screen "BC Process Times" 1280x800, template "Template"
   on GenerateScreen: "TitleUpdater"()
   Button "HmiScreenItemData_1" at 1,1 size 150x43; TextOn 'Back'; TextOff 'Commissioning'
      on Release: ActivateScreen("Commissioning Main Page", 0)
   Button "Button_1" at 21,736 size 161x32; TextOff 'IGG Step Times'
      on Activate: ActivateScreen("IGG Max Step Times", 0)
   Button "Button_2" at 1091,736 size 161x32; TextOff 'BC Step Times'
      on Activate: ActivateScreen("BC Max Step Times", 0)
   AlarmView "Alarm view_1" at 0,777 size 1280x23
   TextField "Text field_2" at 262,326 size 271x22; Text 'CV114 Open Delay Time'
   TextField "Text field_3" at 551,161 size 65x20; Text 'Time (s)'
   TextField "Text field_4" at 262,354 size 273x22; Text 'CV206 Open Delay Time'
   IOField "I/O field_1" at 546,354 size 60x22; Authorization "Parameter Change"; FormatPattern 999
      ProcessValue <- "86_Times_CV206_OPEN_TIME"
   TextField "Text field_5" at 262,411 size 270x22; Text 'CV215 Open Delay Time'
   TextField "Text field_6" at 262,186 size 272x22; Text 'CV127 Open #1 Delay Time'
   TextField "Text field_7" at 262,214 size 272x22; Text 'CV127 Closed Delay Time'
   TextField "Text field_8" at 262,242 size 271x22; Text 'CV127 Open #2 Delay Time'
   TextField "Text field_9" at 262,270 size 270x22; Text 'CV124 Open Delay Time'
   TextField "Text field_10" at 262,298 size 270x22; Text 'CV124 Close Delay Purge Time'
   TextField "Text field_11" at 262,161 size 89x20; Text 'Description'
   IOField "I/O field_3" at 546,186 size 60x22; Authorization "Parameter Change"; FormatPattern 999
      ProcessValue <- "86_Times_CV127_OPEN_TIME_#1"
   IOField "I/O field_4" at 546,214 size 60x22; Authorization "Parameter Change"; FormatPattern 999
      ProcessValue <- "86_Times_CV127_CLOSED_TIME"
   IOField "I/O field_6" at 546,242 size 60x22; Authorization "Parameter Change"; FormatPattern 999
      ProcessValue <- "86_Times_CV127_OPEN_TIME_#2"
   IOField "I/O field_8" at 546,298 size 60x22; Authorization "Parameter Change"; FormatPattern 999
      ProcessValue <- "86_Times_CV124_CLOSE_TIME_PRG"
   IOField "I/O field_9" at 546,410 size 60x22; Authorization "Parameter Change"; FormatPattern 999
      ProcessValue <- "86_Times_CV215_OPEN_TIME"
   TextField "Text field_12" at 261,135 size 178x26; Text 'BC Process Times'
   IOField "I/O field_10" at 546,270 size 60x22; Authorization "Parameter Change"; FormatPattern 999
      ProcessValue <- "86_Times_CV124_OPEN_TIME"
   TextField "Text field_13" at 262,383 size 270x22; Text 'CV207 Open Delay Time'
   IOField "I/O field_11" at 546,382 size 60x22; Authorization "Parameter Change"; FormatPattern 999
      ProcessValue <- "86_Times_CV207_OPEN_TIME"
   TextField "Text field_17" at 262,439 size 270x22; Text 'CV215 Close Delay Purge Time'
   IOField "I/O field_16" at 546,438 size 60x22; Authorization "Parameter Change"; FormatPattern 999
      ProcessValue <- "86_Times_CV215_CLOSE_TIME_PRG"
   TextField "Text field_18" at 262,467 size 270x22; Text 'CV216 Open Delay Time'
   IOField "I/O field_17" at 546,466 size 60x22; Authorization "Parameter Change"; FormatPattern 999
      ProcessValue <- "86_Times_CV216_OPEN_TIME"
   TextField "Text field_19" at 262,495 size 269x22; Text 'CV216 Close Delay Purge Time'
   IOField "I/O field_18" at 546,494 size 60x22; Authorization "Parameter Change"; FormatPattern 999
      ProcessValue <- "86_Times_CV216_CLOSE_TIME_PRG"
   TextField "Text field_20" at 262,523 size 269x22; Text 'CV216 Open Delay Purge Time'
   IOField "I/O field_19" at 546,522 size 60x22; Authorization "Parameter Change"; FormatPattern 999
      ProcessValue <- "86_Times_CV216_OPEN_TIME_PRG"
   TextField "Text field_21" at 262,552 size 269x22; Text 'CV206 Close Delay Time'
   IOField "I/O field_20" at 546,551 size 60x22; Authorization "Parameter Change"; FormatPattern 999
      ProcessValue <- "86_Times_CV206_CLOSE_TIME"
   TextField "Text field_22" at 636,186 size 269x22; Text 'CV207 Close Delay Time'
   IOField "I/O field_21" at 916,186 size 60x22; Authorization "Parameter Change"; FormatPattern 999
      ProcessValue <- "86_Times_CV207_CLOSE_TIME"
   TextField "Text field_23" at 636,160 size 89x20; Text 'Description'
   TextField "Text field_24" at 923,161 size 65x20; Text 'Time (s)'
   TextField "Text field_26" at 636,214 size 269x22; Text 'CV114 Close Delay Time'
   IOField "I/O field_22" at 916,214 size 60x22; Authorization "Parameter Change"; FormatPattern 999
      ProcessValue <- "86_Times_CV114_CLOSE_TIME"
   TextField "Text field_27" at 636,242 size 269x22; Text 'CV215 Close Delay Time'
   IOField "I/O field_23" at 916,242 size 60x22; Authorization "Parameter Change"; FormatPattern 999
      ProcessValue <- "86_Times_CV215_CLOSE_TIME"
   TextField "Text field_28" at 636,270 size 269x22; Text 'CV216 Close Delay Time'
   IOField "I/O field_24" at 916,270 size 60x22; Authorization "Parameter Change"; FormatPattern 999
      ProcessValue <- "86_Times_CV216_CLOSE_TIME"
   TextField "Text field_30" at 636,298 size 269x22; Text 'CV124 Close Delay Time'
   IOField "I/O field_25" at 916,298 size 60x22; Authorization "Parameter Change"; FormatPattern 999
      ProcessValue <- "86_Times_CV124_CLOSE_TIME"
   TextField "Text field_31" at 636,326 size 269x22; Text 'X001 Maximum Run Time'
   IOField "I/O field_26" at 916,326 size 60x22; Authorization "Parameter Change"; FormatPattern 999
      ProcessValue <- "86_Times_X001_MAX_RUN_TIME"
   TextField "Text field_32" at 636,354 size 269x22; Text 'X001 Run Confirmation Time'
   IOField "I/O field_27" at 916,354 size 60x22; Authorization "Parameter Change"; FormatPattern 999
      ProcessValue <- "86_Times_X001_RUN_CNF_TIME"
   TextField "Text field_34" at 636,383 size 269x22; Text 'Flame Detection Delay'
   IOField "I/O field_28" at 916,382 size 60x22; Authorization "Parameter Change"; FormatPattern 999
      ProcessValue <- "86_Times_FD_DET_DELAY"
   TextField "Text field_36" at 636,411 size 269x22; Text 'Flame Verification Time'
   IOField "I/O field_29" at 916,410 size 60x22; Authorization "Parameter Change"; FormatPattern 999
      ProcessValue <- "86_Times_FD_VRFCTN_TIME"
   TextField "Text field_37" at 636,439 size 269x22; Text 'Flame Detection Time'
   IOField "I/O field_30" at 916,438 size 60x22; Authorization "Parameter Change"; FormatPattern 999
      ProcessValue <- "86_Times_FDU_DET_TIME"
   TextField "Text field_38" at 636,467 size 269x22; Text 'Max Ignition Sequence Run Time'
   IOField "I/O field_31" at 916,466 size 60x22; Authorization "Parameter Change"; FormatPattern 999
      ProcessValue <- "86_Times_MAX_IGNTN_SEQ_TIME"
   TextField "Text field_39" at 636,495 size 269x22; Text 'Max Main Burner Sequence Run Time'
      Visibility <- "AlwaysTRUE"
   IOField "I/O field_32" at 916,494 size 60x22; Authorization "Parameter Change"; FormatPattern 999; Unit h
      Visibility <- "AlwaysTRUE"
      ProcessValue <- "86_Times_MAX_MAIN_BURN_SEQ_TIME"
   TextField "Text field_40" at 636,523 size 269x22; Text 'Max Pilot Burner Purge Sequence Run Time'
   IOField "I/O field_33" at 916,522 size 60x22; Authorization "Parameter Change"; FormatPattern 999
      ProcessValue <- "86_Times_MAX_PILOT_PURGE_SEQ_TIME"
   TextField "Text field_41" at 636,552 size 269x22; Text 'O2 Check Delay Time'
   IOField "I/O field_34" at 916,551 size 60x22; Authorization "Parameter Change"; FormatPattern 999
      ProcessValue <- "86_Times_O2_CHECK_TIME"
   IOField "I/O field_7" at 546,326 size 60x22; Authorization "Parameter Change"; FormatPattern 999
      ProcessValue <- "86_Times_CV114_OPEN_TIME"
   TextField "Text field_43" at 636,582 size 269x22; Text 'Flame Fail Delay'
   IOField "I/O field_35" at 916,581 size 60x22; Authorization "Parameter Change"; FormatPattern 999
      ProcessValue <- "80_From_HMI_FLM_FAIL_DLY"
   Switch "Switch_1" at 987,492 size 32x29; CaptionText 'Switch'; TextOn 'ON'; TextOff 'OFF'; Authorization "User administration"; PictureOff "Design_5_PilotLight_Green_Off"; PictureOn "Design_5_PilotLight_Green_On"
      on Activate: SetBit("80_From_HMI_BurnerProgramedStop")
      Visibility <- "AlwaysTRUE"
      ProcessValue <- "80_From_HMI_BurnerProgramedStop"
   TextField "Text field_44" at 636,613 size 269x22; Text 'FS317 Delayed Fault'
   IOField "I/O field_36" at 916,613 size 60x22; Authorization "Parameter Change"; FormatPattern 999
      ProcessValue <- "86_Times_FS317 delay"
   TextField "Text field_45" at 636,644 size 269x22; Text 'FS320 Delayed Fault'
   IOField "I/O field_37" at 916,644 size 60x22; Authorization "Parameter Change"; FormatPattern 999
      ProcessValue <- "86_Times_FS320 delay"
   TextField "Text field_46" at 262,581 size 269x22; Text 'FS359 Delayed Fault'
   IOField "I/O field_38" at 546,581 size 60x22; Authorization "Parameter Change"; FormatPattern 999
      ProcessValue <- "80_From_HMI_PIT 359 delay"
   TextField "Text field_47" at 262,612 size 269x22; Text 'FS316 Delayed Fault'
   IOField "I/O field_39" at 546,612 size 60x22; Authorization "Parameter Change"; FormatPattern 999
      ProcessValue <- "80_From_HMI_PIT 316 delay"
   Group "Group" at 455,41 size 373x50
   TextField "Text field_1" at 262,643 size 269x22; Text 'PS101 Delayed Fault'
   IOField "I/O field_2" at 546,643 size 60x22; Authorization "Parameter Change"; FormatPattern 999
      ProcessValue <- "86_Times_PS101 Alarm Delay"
   Button "HmiScreenItemData_8" at 469,45 size 355x40; TextOn 'Back'; TextOff 'Text'
   TextField "Screen title" at 455,41 size 373x50; Text 'Screen title'

screen "GCU Process Times" 1280x800, template "Template"
   on GenerateScreen: "TitleUpdater"()
   Button "HmiScreenItemData_1" at 1,1 size 150x43; TextOn 'Back'; TextOff 'Commissioning'
      on Release: ActivateScreen("Commissioning Main Page", 0)
   AlarmView "Alarm view_1" at 0,777 size 1280x23
   TextField "Text field_29" at 545,103 size 65x20; Text 'Time (s)'
   TextField "Text field_65" at 240,128 size 300x25; Text 'P303 Started Delay'
   TextField "Text field_42" at 240,103 size 89x20; Text 'Description'
   IOField "I/O field_128" at 545,128 size 65x25; Authorization "Parameter Change"; FormatPattern 999
      ProcessValue <- "86_Times_P303_STRTD_DLY"
   TextField "Text field_53" at 240,74 size 193x26; Text 'GCU Process Times'
   TextField "Text field_1" at 240,158 size 300x25; Text 'P303 Stopped Delay'
   IOField "I/O field_1" at 545,158 size 65x25; Authorization "Parameter Change"; FormatPattern 999
      ProcessValue <- "86_Times_P303_STPD_DLY"
   TextField "Text field_2" at 240,188 size 300x25; Text 'P304 Started Delay'
   IOField "I/O field_2" at 545,188 size 65x25; Authorization "Parameter Change"; FormatPattern 999
      ProcessValue <- "86_Times_P304_STRTD_DLY"
   TextField "Text field_3" at 240,218 size 300x25; Text 'P304 Stopped Delay'
   IOField "I/O field_3" at 545,218 size 65x25; Authorization "Parameter Change"; FormatPattern 999
      ProcessValue <- "86_Times_P304_STPD_DLY"
   TextField "Text field_4" at 240,248 size 300x25; Text 'P305 Started Delay'
   IOField "I/O field_4" at 545,248 size 65x25; Authorization "Parameter Change"; FormatPattern 999
      ProcessValue <- "86_Times_P305_STRTD_DLY"
   TextField "Text field_5" at 240,278 size 300x25; Text 'P305 Stopped Delay'
   IOField "I/O field_5" at 545,278 size 65x25; Authorization "Parameter Change"; FormatPattern 999
      ProcessValue <- "86_Times_P305_STPD_DLY"
   TextField "Text field_6" at 240,308 size 300x25; Text 'CV341 Closed Delay'
   IOField "I/O field_6" at 545,308 size 65x25; Authorization "Parameter Change"; FormatPattern 999
      ProcessValue <- "86_Times_CV341_CLSD_DLY"
   TextField "Text field_7" at 240,338 size 300x25; Text 'CV358 Closed Delay'
   IOField "I/O field_7" at 545,338 size 65x25; Authorization "Parameter Change"; FormatPattern 999
      ProcessValue <- "86_Times_CV358_CLSD_DLY"
   TextField "Text field_8" at 975,103 size 65x20; Text 'Time (s)'
   TextField "Text field_9" at 670,128 size 300x25; Text 'CV405 Opened Delay'
   TextField "Text field_10" at 670,103 size 89x20; Text 'Description'
   IOField "I/O field_8" at 975,128 size 65x25; Authorization "Parameter Change"; FormatPattern 999
      ProcessValue <- "86_Times_CV405_OPND_DLY"
   TextField "Text field_11" at 670,158 size 300x25; Text 'CV406 Closed Delay'
   IOField "I/O field_9" at 975,158 size 65x25; Authorization "Parameter Change"; FormatPattern 999
      ProcessValue <- "86_Times_CV406_CLSD_DLY"
   TextField "Text field_12" at 670,188 size 300x25; Text 'E400 Stop Time'
   IOField "I/O field_10" at 975,188 size 65x25; Authorization "Parameter Change"; FormatPattern 999
      ProcessValue <- "86_Times_E400_STOP_TIME"
   TextField "Text field_13" at 670,218 size 300x25; Text 'P303 Stop Time'
   IOField "I/O field_11" at 975,218 size 65x25; Authorization "Parameter Change"; FormatPattern 999
      ProcessValue <- "86_Times_P303_STOP_TIME"
   TextField "Text field_14" at 670,248 size 300x25; Text 'CV341 Opened Delay'
   IOField "I/O field_12" at 975,248 size 65x25; Authorization "Parameter Change"; FormatPattern 999
      ProcessValue <- "86_Times_CV341_OPND_DLY"
   TextField "Text field_15" at 670,278 size 300x25; Text 'GCU Tank Maximum Drain Time'
   IOField "I/O field_13" at 975,278 size 65x25; Authorization "Parameter Change"; FormatPattern 999
      ProcessValue <- "86_Times_GCU_TNK_DRN_MAX_TIME"
   TextField "Text field_16" at 670,308 size 300x25; Text 'GCU Flush Time'
   IOField "I/O field_14" at 975,308 size 65x25; Authorization "Parameter Change"; FormatPattern 999
      ProcessValue <- "86_Times_GCU_FLUSH_TIME"
   TextField "Text field_17" at 670,338 size 300x25; Text 'Post Flush Delay'
   IOField "I/O field_15" at 975,338 size 65x25; Authorization "Parameter Change"; FormatPattern 999
      ProcessValue <- "86_Times_POST_FLUSH_DLY"
   TextField "Text field_18" at 240,368 size 300x25; Text 'CV401 Opened Delay'
   IOField "I/O field_16" at 545,368 size 65x25; Authorization "Parameter Change"; FormatPattern 999
      ProcessValue <- "86_Times_CV401_OPND_DLY"
   TextField "Text field_19" at 240,398 size 300x25; Text 'CV401 Closed Delay'
   IOField "I/O field_17" at 545,398 size 65x25; Authorization "Parameter Change"; FormatPattern 999
      ProcessValue <- "86_Times_CV401_CLSD_DLY"
   TextField "Text field_20" at 240,428 size 300x25; Text 'CV441 Opened Delay'
   IOField "I/O field_18" at 545,428 size 65x25; Authorization "Parameter Change"; FormatPattern 999
      ProcessValue <- "86_Times_CV441_OPND_DLY"
   TextField "Text field_21" at 240,458 size 300x25; Text 'CV441 Closed Delay'
   IOField "I/O field_19" at 545,458 size 65x25; Authorization "Parameter Change"; FormatPattern 999
      ProcessValue <- "86_Times_CV441_CLSD_DLY"
   TextField "Text field_22" at 240,488 size 300x25; Text 'Pre CV441 Open Delay'
   IOField "I/O field_20" at 545,488 size 65x25; Authorization "Parameter Change"; FormatPattern 999
      ProcessValue <- "86_Times_PRE_CV441_OPN_DLY"
   TextField "Text field_23" at 240,518 size 300x25; Text 'Valve Configuration Done Delay'
   IOField "I/O field_21" at 545,518 size 65x25; Authorization "Parameter Change"; FormatPattern 999
      ProcessValue <- "86_Times_VLV_CNFG_DN_DLY"
   TextField "Text field_24" at 240,548 size 300x25; Text 'Pre GCU Tank Fill Delay'
   IOField "I/O field_22" at 545,548 size 65x25; Authorization "Parameter Change"; FormatPattern 999
      ProcessValue <- "86_Times_PRE_GCU_TNK_FILL_DLY"
   TextField "Text field_25" at 240,578 size 300x25; Text 'GCU Tank Fill Maximum Time'
   IOField "I/O field_23" at 545,578 size 65x25; Authorization "Parameter Change"; FormatPattern 999
      ProcessValue <- "86_Times_GCU_TNK_FILL_MAX_TIME"
   TextField "Text field_26" at 670,368 size 300x25; Text 'CV341 Maximum Travel Time'
   IOField "I/O field_24" at 975,368 size 65x25; Authorization "Parameter Change"; FormatPattern 999
      ProcessValue <- "86_Times_CV341_MAX_TRVL_TIME"
   TextField "Text field_27" at 670,398 size 300x25; Text 'CV358 Maximum Travel Time'
   IOField "I/O field_25" at 975,398 size 65x25; Authorization "Parameter Change"; FormatPattern 999
      ProcessValue <- "86_Times_CV358_MAX_TRVL_TIME"
   TextField "Text field_28" at 670,428 size 300x25; Text 'CV406 Maximum Travel Time'
   IOField "I/O field_26" at 975,428 size 65x25; Authorization "Parameter Change"; FormatPattern 999
      ProcessValue <- "86_Times_CV406_MAX_TRVL_TIME"
   TextField "Text field_30" at 670,458 size 300x25; Text 'CV407 Maximum Travel Time'
   IOField "I/O field_27" at 975,458 size 65x25; Authorization "Parameter Change"; FormatPattern 999
      ProcessValue <- "86_Times_CV407_MAX_TRVL_TIME"
   TextField "Text field_31" at 670,488 size 300x25; Text 'CV409 Maximum Travel Time'
   IOField "I/O field_28" at 975,488 size 65x25; Authorization "Parameter Change"; FormatPattern 999
      ProcessValue <- "86_Times_CV409_MAX_TRVL_TIME"
   TextField "Text field_32" at 670,518 size 300x25; Text 'CV411 Maximum Travel Time'
   IOField "I/O field_29" at 975,518 size 65x25; Authorization "Parameter Change"; FormatPattern 999
      ProcessValue <- "86_Times_CV411_MAX_TRVL_TIME"
   TextField "Text field_33" at 670,548 size 300x25; Text 'CV441 Maximum Travel Time'
   IOField "I/O field_30" at 975,548 size 65x25; Authorization "Parameter Change"; FormatPattern 999
      ProcessValue <- "86_Times_CV441_MAX_TRVL_TIME"
   TextField "Text field_34" at 670,638 size 300x25; Text 'PIT416 Target Ramp Time'
   IOField "I/O field_31" at 975,638 size 65x25; Authorization "Parameter Change"; FormatPattern 999
      ProcessValue <- "86_Times_PIT416_TRGT_RMP_TIME"
   TextField "Text field_35" at 240,608 size 300x25; Text 'E400 Started Delay'
   IOField "I/O field_32" at 545,608 size 65x25; Authorization "Parameter Change"; FormatPattern 999
      ProcessValue <- "86_Times_E400_STRTD_DLY"
   TextField "Text field_36" at 240,638 size 300x25; Text 'E400 Running Delay'
   IOField "I/O field_33" at 545,638 size 65x25; Authorization "Parameter Change"; FormatPattern 999
      ProcessValue <- "86_Times_E400_RNG_DLY"
   TextField "Text field_37" at 670,578 size 300x25; Text 'PIT353 Alarm Delay Time'
   IOField "I/O field_34" at 975,578 size 65x25; Authorization "Parameter Change"; FormatPattern 999
      ProcessValue <- "86_Times_PIT353 Delay"
   TextField "Text field_38" at 670,608 size 300x25; Text 'PIT416 Alarm Delay Time'
   IOField "I/O field_35" at 975,608 size 65x25; Authorization "Parameter Change"; FormatPattern 999
      ProcessValue <- "86_Times_PIT416 Delay"
   TextField "Text field_39" at 240,669 size 300x25; Text 'P301 Started Delay'
   IOField "I/O field_36" at 545,669 size 65x25; Authorization "Parameter Change"; FormatPattern 999
      ProcessValue <- "86_Times_P301_START_DLY"
   TextField "Text field_40" at 670,669 size 300x25; Text 'FS332 Alarm Delay'
   IOField "I/O field_37" at 975,669 size 65x25; Authorization "Parameter Change"; FormatPattern 999
      ProcessValue <- "86_Times_FS332 Delay"
   TextField "Text field_41" at 670,701 size 300x25; Text 'LIT304 Alarm Delay'
   IOField "I/O field_38" at 975,701 size 65x25; Authorization "Parameter Change"; FormatPattern 999
      ProcessValue <- "86_Times_LIT304 Delay"
   Group "Group" at 455,41 size 373x50
   TextField "Text field_43" at 240,701 size 300x25; Text 'PIT358 Alarm Delay Time'
   IOField "I/O field_39" at 545,701 size 65x25; Authorization "Parameter Change"; FormatPattern 999
      ProcessValue <- "86_Times_PIT358 Delay"
   TextField "Text field_44" at 240,732 size 300x25; Text 'PIT348 Alarm Delay Time'
   IOField "I/O field_40" at 545,732 size 65x25; Authorization "Parameter Change"; FormatPattern 999
      ProcessValue <- "86_Times_PIT348 Delay"
   Button "HmiScreenItemData_8" at 469,45 size 355x40; TextOn 'Back'; TextOff 'Text'
   TextField "Screen title" at 455,41 size 373x50; Text 'Screen title'

screen "GCU Max Step Times" 1280x800, template "Template"
   on GenerateScreen: "TitleUpdater"()
   Button "HmiScreenItemData_1" at 1,1 size 150x43; TextOn 'Back'; TextOff 'Commissioning'
      on Release: ActivateScreen("Commissioning Main Page", 0)
   TextField "Text field_29" at 130,95 size 75x25; Text 'Time (ms)'
   TextField "Text field_65" at 40,130 size 75x25; Text 'Step 001'
   TextField "Text field_42" at 40,95 size 75x25; Text 'STEP'
   IOField "I/O field_128" at 130,130 size 75x25; Authorization "Parameter Change"; FormatPattern 999999
      ProcessValue <- "86_Times_STEP_MAX_TIME_STP_001"
   TextField "Text field_53" at 40,66 size 262x26; Text 'GCU Maximum Step Times'
   TextField "Text field_1" at 385,95 size 75x25; Text 'Time (ms)'
   TextField "Text field_2" at 295,130 size 75x25; Text 'Step 170'
   TextField "Text field_3" at 295,95 size 75x25; Text 'STEP'
   IOField "I/O field_1" at 385,130 size 75x25; Authorization "Parameter Change"; FormatPattern 999999
      ProcessValue <- "86_Times_STEP_MAX_TIME_STP_170"
   TextField "Text field_4" at 640,95 size 75x25; Text 'Time (ms)'
   TextField "Text field_5" at 550,130 size 75x25; Text 'Step 350'
   TextField "Text field_6" at 550,95 size 75x25; Text 'STEP'
   IOField "I/O field_2" at 640,130 size 75x25; Authorization "Parameter Change"; FormatPattern 999999
      ProcessValue <- "86_Times_STEP_MAX_TIME_STP_350"
   TextField "Text field_7" at 895,95 size 75x25; Text 'Time (ms)'
   TextField "Text field_8" at 805,130 size 75x25; Text 'Step 530'
   TextField "Text field_9" at 805,95 size 75x25; Text 'STEP'
   IOField "I/O field_3" at 895,130 size 75x25; Authorization "Parameter Change"; FormatPattern 999999
      ProcessValue <- "86_Times_STEP_MAX_TIME_STP_530"
   TextField "Text field_10" at 1150,95 size 75x25; Text 'Time (ms)'
   TextField "Text field_12" at 1060,95 size 75x25; Text 'STEP'
   TextField "Text field_13" at 40,165 size 75x25; Text 'Step 005'
   IOField "I/O field_5" at 130,165 size 75x25; Authorization "Parameter Change"; FormatPattern 999999
      ProcessValue <- "86_Times_STEP_MAX_TIME_STP_005"
   TextField "Text field_14" at 295,165 size 75x25; Text 'Step 180'
   IOField "I/O field_6" at 385,165 size 75x25; Authorization "Parameter Change"; FormatPattern 999999
      ProcessValue <- "86_Times_STEP_MAX_TIME_STP_180"
   TextField "Text field_15" at 550,165 size 75x25; Text 'Step 360'
   IOField "I/O field_7" at 640,165 size 75x25; Authorization "Parameter Change"; FormatPattern 999999
      ProcessValue <- "86_Times_STEP_MAX_TIME_STP_360"
   TextField "Text field_16" at 805,165 size 75x25; Text 'Step 540'
   IOField "I/O field_8" at 895,165 size 75x25; Authorization "Parameter Change"; FormatPattern 999999
      ProcessValue <- "86_Times_STEP_MAX_TIME_STP_540"
   TextField "Text field_18" at 40,200 size 75x25; Text 'Step 010'
   IOField "I/O field_10" at 130,200 size 75x25; Authorization "Parameter Change"; FormatPattern 999999
      ProcessValue <- "86_Times_STEP_MAX_TIME_STP_010"
   TextField "Text field_19" at 295,200 size 75x25; Text 'Step 190'
   IOField "I/O field_11" at 385,200 size 75x25; Authorization "Parameter Change"; FormatPattern 999999
      ProcessValue <- "86_Times_STEP_MAX_TIME_STP_190"
   TextField "Text field_20" at 550,200 size 75x25; Text 'Step 370'
   IOField "I/O field_12" at 640,200 size 75x25; Authorization "Parameter Change"; FormatPattern 999999
      ProcessValue <- "86_Times_STEP_MAX_TIME_STP_370"
   TextField "Text field_21" at 805,200 size 75x25; Text 'Step 550'
   IOField "I/O field_13" at 895,200 size 75x25; Authorization "Parameter Change"; FormatPattern 999999
      ProcessValue <- "86_Times_STEP_MAX_TIME_STP_550"
   TextField "Text field_23" at 40,235 size 75x25; Text 'Step 020'
   IOField "I/O field_15" at 130,235 size 75x25; Authorization "Parameter Change"; FormatPattern 999999
      ProcessValue <- "86_Times_STEP_MAX_TIME_STP_020"
   TextField "Text field_24" at 295,235 size 75x25; Text 'Step 200'
   IOField "I/O field_16" at 385,235 size 75x25; Authorization "Parameter Change"; FormatPattern 999999
      ProcessValue <- "86_Times_STEP_MAX_TIME_STP_200"
   TextField "Text field_25" at 550,235 size 75x25; Text 'Step 380'
   IOField "I/O field_17" at 640,235 size 75x25; Authorization "Parameter Change"; FormatPattern 999999
      ProcessValue <- "86_Times_STEP_MAX_TIME_STP_380"
   TextField "Text field_26" at 805,235 size 75x25; Text 'Step 560'
   IOField "I/O field_18" at 895,235 size 75x25; Authorization "Parameter Change"; FormatPattern 999999
      ProcessValue <- "86_Times_STEP_MAX_TIME_STP_560"
   TextField "Text field_28" at 40,270 size 75x25; Text 'Step 030'
   IOField "I/O field_20" at 130,270 size 75x25; Authorization "Parameter Change"; FormatPattern 999999
      ProcessValue <- "86_Times_STEP_MAX_TIME_STP_030"
   TextField "Text field_30" at 295,270 size 75x25; Text 'Step 210'
   IOField "I/O field_21" at 385,270 size 75x25; Authorization "Parameter Change"; FormatPattern 999999
      ProcessValue <- "86_Times_STEP_MAX_TIME_STP_210"
   TextField "Text field_31" at 550,270 size 75x25; Text 'Step 390'
   IOField "I/O field_22" at 640,270 size 75x25; Authorization "Parameter Change"; FormatPattern 999999
      ProcessValue <- "86_Times_STEP_MAX_TIME_STP_390"
   TextField "Text field_32" at 805,270 size 75x25; Text 'Step 570'
   IOField "I/O field_23" at 895,270 size 75x25; Authorization "Parameter Change"; FormatPattern 999999
      ProcessValue <- "86_Times_STEP_MAX_TIME_STP_570"
   TextField "Text field_34" at 40,305 size 75x25; Text 'Step 040'
   IOField "I/O field_25" at 130,305 size 75x25; Authorization "Parameter Change"; FormatPattern 999999
      ProcessValue <- "86_Times_STEP_MAX_TIME_STP_040"
   TextField "Text field_35" at 295,305 size 75x25; Text 'Step 220'
   IOField "I/O field_26" at 385,305 size 75x25; Authorization "Parameter Change"; FormatPattern 999999
      ProcessValue <- "86_Times_STEP_MAX_TIME_STP_220"
   TextField "Text field_36" at 550,305 size 75x25; Text 'Step 400'
   IOField "I/O field_27" at 640,305 size 75x25; Authorization "Parameter Change"; FormatPattern 999999
      ProcessValue <- "86_Times_STEP_MAX_TIME_STP_400"
   TextField "Text field_37" at 805,305 size 75x25; Text 'Step 580'
   IOField "I/O field_28" at 895,305 size 75x25; Authorization "Parameter Change"; FormatPattern 999999
      ProcessValue <- "86_Times_STEP_MAX_TIME_STP_580"
   TextField "Text field_39" at 40,340 size 75x25; Text 'Step 050'
   IOField "I/O field_30" at 130,340 size 75x25; Authorization "Parameter Change"; FormatPattern 999999
      ProcessValue <- "86_Times_STEP_MAX_TIME_STP_050"
   TextField "Text field_40" at 295,340 size 75x25; Text 'Step 230'
   IOField "I/O field_31" at 385,340 size 75x25; Authorization "Parameter Change"; FormatPattern 999999
      ProcessValue <- "86_Times_STEP_MAX_TIME_STP_230"
   TextField "Text field_41" at 550,340 size 75x25; Text 'Step 410'
   IOField "I/O field_32" at 640,340 size 75x25; Authorization "Parameter Change"; FormatPattern 999999
      ProcessValue <- "86_Times_STEP_MAX_TIME_STP_410"
   TextField "Text field_43" at 805,340 size 75x25; Text 'Step 590'
   IOField "I/O field_33" at 895,340 size 75x25; Authorization "Parameter Change"; FormatPattern 999999
      ProcessValue <- "86_Times_STEP_MAX_TIME_STP_590"
   TextField "Text field_45" at 40,375 size 75x25; Text 'Step 060'
   IOField "I/O field_35" at 130,375 size 75x25; Authorization "Parameter Change"; FormatPattern 999999
      ProcessValue <- "86_Times_STEP_MAX_TIME_STP_060"
   TextField "Text field_46" at 295,375 size 75x25; Text 'Step 240'
   IOField "I/O field_36" at 385,375 size 75x25; Authorization "Parameter Change"; FormatPattern 999999
      ProcessValue <- "86_Times_STEP_MAX_TIME_STP_240"
   TextField "Text field_47" at 550,375 size 75x25; Text 'Step 420'
   IOField "I/O field_37" at 640,375 size 75x25; Authorization "Parameter Change"; FormatPattern 999999
      ProcessValue <- "86_Times_STEP_MAX_TIME_STP_420"
   TextField "Text field_48" at 805,375 size 75x25; Text 'Step 600'
   IOField "I/O field_38" at 895,375 size 75x25; Authorization "Parameter Change"; FormatPattern 999999
      ProcessValue <- "86_Times_STEP_MAX_TIME_STP_600"
   TextField "Text field_50" at 40,410 size 75x25; Text 'Step 070'
   IOField "I/O field_40" at 130,410 size 75x25; Authorization "Parameter Change"; FormatPattern 999999
      ProcessValue <- "86_Times_STEP_MAX_TIME_STP_070"
   TextField "Text field_51" at 295,410 size 75x25; Text 'Step 250'
   IOField "I/O field_41" at 385,410 size 75x25; Authorization "Parameter Change"; FormatPattern 999999
      ProcessValue <- "86_Times_STEP_MAX_TIME_STP_250"
   TextField "Text field_52" at 550,410 size 75x25; Text 'Step 430'
   IOField "I/O field_42" at 640,410 size 75x25; Authorization "Parameter Change"; FormatPattern 999999
      ProcessValue <- "86_Times_STEP_MAX_TIME_STP_430"
   TextField "Text field_54" at 805,410 size 75x25; Text 'Step 610'
   IOField "I/O field_43" at 895,410 size 75x25; Authorization "Parameter Change"; FormatPattern 999999
      ProcessValue <- "86_Times_STEP_MAX_TIME_STP_610"
   TextField "Text field_56" at 40,445 size 75x25; Text 'Step 080'
   IOField "I/O field_45" at 130,445 size 75x25; Authorization "Parameter Change"; FormatPattern 999999
      ProcessValue <- "86_Times_STEP_MAX_TIME_STP_080"
   TextField "Text field_57" at 295,445 size 75x25; Text 'Step 260'
   IOField "I/O field_46" at 385,445 size 75x25; Authorization "Parameter Change"; FormatPattern 999999
      ProcessValue <- "86_Times_STEP_MAX_TIME_STP_260"
   TextField "Text field_58" at 550,445 size 75x25; Text 'Step 440'
   IOField "I/O field_47" at 640,445 size 75x25; Authorization "Parameter Change"; FormatPattern 999999
      ProcessValue <- "86_Times_STEP_MAX_TIME_STP_440"
   TextField "Text field_59" at 805,445 size 75x25; Text 'Step 620'
   IOField "I/O field_48" at 895,445 size 75x25; Authorization "Parameter Change"; FormatPattern 999999
      ProcessValue <- "86_Times_STEP_MAX_TIME_STP_620"
   TextField "Text field_61" at 40,480 size 75x25; Text 'Step 090'
   IOField "I/O field_50" at 130,480 size 75x25; Authorization "Parameter Change"; FormatPattern 999999
      ProcessValue <- "86_Times_STEP_MAX_TIME_STP_090"
   TextField "Text field_62" at 295,480 size 75x25; Text 'Step 270'
   IOField "I/O field_51" at 385,480 size 75x25; Authorization "Parameter Change"; FormatPattern 999999
      ProcessValue <- "86_Times_STEP_MAX_TIME_STP_270"
   TextField "Text field_63" at 550,480 size 75x25; Text 'Step 450'
   IOField "I/O field_52" at 640,480 size 75x25; Authorization "Parameter Change"; FormatPattern 999999
      ProcessValue <- "86_Times_STEP_MAX_TIME_STP_450"
   TextField "Text field_64" at 805,480 size 75x25; Text 'Step 630'
   IOField "I/O field_53" at 895,480 size 75x25; Authorization "Parameter Change"; FormatPattern 999999
      ProcessValue <- "86_Times_STEP_MAX_TIME_STP_630"
   TextField "Text field_67" at 40,515 size 75x25; Text 'Step 100'
   IOField "I/O field_55" at 130,515 size 75x25; Authorization "Parameter Change"; FormatPattern 999999
      ProcessValue <- "86_Times_STEP_MAX_TIME_STP_100"
   TextField "Text field_68" at 295,515 size 75x25; Text 'Step 280'
   IOField "I/O field_56" at 385,515 size 75x25; Authorization "Parameter Change"; FormatPattern 999999
      ProcessValue <- "86_Times_STEP_MAX_TIME_STP_280"
   TextField "Text field_69" at 550,515 size 75x25; Text 'Step 460'
   IOField "I/O field_57" at 640,515 size 75x25; Authorization "Parameter Change"; FormatPattern 999999
      ProcessValue <- "86_Times_STEP_MAX_TIME_STP_460"
   TextField "Text field_72" at 40,550 size 75x25; Text 'Step 110'
   IOField "I/O field_60" at 130,550 size 75x25; Authorization "Parameter Change"; FormatPattern 999999
      ProcessValue <- "86_Times_STEP_MAX_TIME_STP_110"
   TextField "Text field_73" at 295,550 size 75x25; Text 'Step 290'
   IOField "I/O field_61" at 385,550 size 75x25; Authorization "Parameter Change"; FormatPattern 999999
      ProcessValue <- "86_Times_STEP_MAX_TIME_STP_290"
   TextField "Text field_74" at 550,550 size 75x25; Text 'Step 470'
   IOField "I/O field_62" at 640,550 size 75x25; Authorization "Parameter Change"; FormatPattern 999999
      ProcessValue <- "86_Times_STEP_MAX_TIME_STP_470"
   TextField "Text field_77" at 40,585 size 75x25; Text 'Step 120'
   IOField "I/O field_65" at 130,585 size 75x25; Authorization "Parameter Change"; FormatPattern 999999
      ProcessValue <- "86_Times_STEP_MAX_TIME_STP_120"
   TextField "Text field_78" at 295,585 size 75x25; Text 'Step 300'
   IOField "I/O field_66" at 385,585 size 75x25; Authorization "Parameter Change"; FormatPattern 999999
      ProcessValue <- "86_Times_STEP_MAX_TIME_STP_300"
   TextField "Text field_79" at 550,585 size 75x25; Text 'Step 480'
   IOField "I/O field_67" at 640,585 size 75x25; Authorization "Parameter Change"; FormatPattern 999999
      ProcessValue <- "86_Times_STEP_MAX_TIME_STP_480"
   TextField "Text field_82" at 40,620 size 75x25; Text 'Step 130'
   IOField "I/O field_70" at 130,620 size 75x25; Authorization "Parameter Change"; FormatPattern 999999
      ProcessValue <- "86_Times_STEP_MAX_TIME_STP_130"
   TextField "Text field_83" at 295,620 size 75x25; Text 'Step 310'
   IOField "I/O field_71" at 385,620 size 75x25; Authorization "Parameter Change"; FormatPattern 999999
      ProcessValue <- "86_Times_STEP_MAX_TIME_STP_310"
   TextField "Text field_84" at 550,620 size 75x25; Text 'Step 490'
   IOField "I/O field_72" at 640,620 size 75x25; Authorization "Parameter Change"; FormatPattern 999999
      ProcessValue <- "86_Times_STEP_MAX_TIME_STP_490"
   TextField "Text field_87" at 40,655 size 75x25; Text 'Step 140'
   IOField "I/O field_75" at 130,655 size 75x25; Authorization "Parameter Change"; FormatPattern 999999
      ProcessValue <- "86_Times_STEP_MAX_TIME_STP_140"
   TextField "Text field_88" at 295,655 size 75x25; Text 'Step 320'
   IOField "I/O field_76" at 385,655 size 75x25; Authorization "Parameter Change"; FormatPattern 999999
      ProcessValue <- "86_Times_STEP_MAX_TIME_STP_320"
   TextField "Text field_89" at 550,655 size 75x25; Text 'Step 500'
   IOField "I/O field_77" at 640,655 size 75x25; Authorization "Parameter Change"; FormatPattern 999999
      ProcessValue <- "86_Times_STEP_MAX_TIME_STP_500"
   TextField "Text field_92" at 40,690 size 75x25; Text 'Step 150'
   IOField "I/O field_80" at 130,690 size 75x25; Authorization "Parameter Change"; FormatPattern 999999
      ProcessValue <- "86_Times_STEP_MAX_TIME_STP_150"
   TextField "Text field_93" at 295,690 size 75x25; Text 'Step 330'
   IOField "I/O field_81" at 385,690 size 75x25; Authorization "Parameter Change"; FormatPattern 999999
      ProcessValue <- "86_Times_STEP_MAX_TIME_STP_330"
   TextField "Text field_94" at 550,690 size 75x25; Text 'Step 510'
   IOField "I/O field_82" at 640,690 size 75x25; Authorization "Parameter Change"; FormatPattern 999999
      ProcessValue <- "86_Times_STEP_MAX_TIME_STP_510"
   TextField "Text field_97" at 40,725 size 75x25; Text 'Step 160'
   IOField "I/O field_85" at 130,725 size 75x25; Authorization "Parameter Change"; FormatPattern 999999
      ProcessValue <- "86_Times_STEP_MAX_TIME_STP_160"
   TextField "Text field_98" at 295,725 size 75x25; Text 'Step 340'
   IOField "I/O field_86" at 385,725 size 75x25; Authorization "Parameter Change"; FormatPattern 999999
      ProcessValue <- "86_Times_STEP_MAX_TIME_STP_340"
   TextField "Text field_99" at 550,725 size 75x25; Text 'Step 520'
   IOField "I/O field_87" at 640,725 size 75x25; Authorization "Parameter Change"; FormatPattern 999999
      ProcessValue <- "86_Times_STEP_MAX_TIME_STP_520"
   Group "Group" at 455,41 size 373x50
   Button "HmiScreenItemData_8" at 469,45 size 355x40; TextOn 'Back'; TextOff 'Text'
   TextField "Screen title" at 455,41 size 373x50; Text 'Screen title'

screen "GCU Target Setpoints" 1280x800, template "Template"
   on GenerateScreen: "TitleUpdater"()
   Button "HmiScreenItemData_1" at 1,1 size 150x43; TextOn 'Back'; TextOff 'Commissioning'
      on Release: ActivateScreen("Commissioning Main Page", 0)
   AlarmView "Alarm view_1" at 0,777 size 1280x23
   TextField "Text field_37" at 20,239 size 300x30; Text 'GCU Control PLC (Rack 3)'
   TextField "Text field_1" at 810,239 size 450x30; Text 'PROCESS STEP RELATED SETPOINTS & TARGETS'
   TextField "Text field_82" at 100,299 size 220x22; Text 'LIT304 GCU LEVEL'
   IOField "I/O field_22" at 350,299 size 70x22; FormatPattern 999; Unit  %
      ProcessValue <- "12_AI_Data_LIT_304_SCALED"
   IOField "I/O field_23" at 450,299 size 75x22; Authorization "Parameter Change"; FormatPattern 999
      ProcessValue <- "84_Setpoints_LIT304_InitialFill_LowLow"
   IOField "I/O field_24" at 550,299 size 75x22; Authorization "Parameter Change"; FormatPattern 999
      ProcessValue <- "84_Setpoints_LIT304_InitialFill_Low"
   IOField "I/O field_25" at 952,299 size 75x22; Authorization "Parameter Change"; FormatPattern 999
      ProcessValue <- "84_Setpoints_LIT304_InitialFill_High"
   IOField "I/O field_26" at 1052,299 size 75x22; Authorization "Parameter Change"; FormatPattern 999
      ProcessValue <- "84_Setpoints_LIT304_InitialFill_HighHigh"
   TextField "Text field_22" at 20,299 size 53x22; Text 'IW800'
   TextField "Text field_90" at 350,272 size 70x22; Text 'Reading'
   TextField "Text field_23" at 450,272 size 75x22; Text 'Low Low'
   TextField "Text field_26" at 550,272 size 75x22; Text 'Low'
   TextField "Text field_27" at 952,272 size 75x22; Text 'High'
   TextField "Text field_28" at 1052,272 size 75x22; Text 'High High'
   TextField "Text field_41" at 100,272 size 220x22; Text 'Description'
   TextField "Text field_43" at 20,272 size 53x22; Text 'AI'
   IOField "I/O field_27" at 750,299 size 75x22; Authorization "Parameter Change"; FormatPattern 999
      ProcessValue <- "84_Setpoints_LIT304_InitialFill_Target"
   TextField "Text field_29" at 750,272 size 75x22; Text 'Target'
   TextField "Text field_30" at 1152,299 size 100x22; Text 'INITIAL FILL'
   IOField "I/O field_28" at 450,339 size 75x22; Authorization "Parameter Change"; FormatPattern 999
      ProcessValue <- "84_Setpoints_LIT304_Refill_LowLow"
   IOField "I/O field_29" at 550,339 size 75x22; Authorization "Parameter Change"; FormatPattern 999
      ProcessValue <- "84_Setpoints_LIT304_Refill_Low"
   IOField "I/O field_30" at 952,339 size 75x22; Authorization "Parameter Change"; FormatPattern 999
      ProcessValue <- "84_Setpoints_LIT304_Refill_High"
   IOField "I/O field_40" at 1052,339 size 75x22; Authorization "Parameter Change"; FormatPattern 999
      ProcessValue <- "84_Setpoints_LIT304_Refill_HighHigh"
   IOField "I/O field_43" at 650,339 size 75x22; Authorization "Parameter Change"; FormatPattern 999
      ProcessValue <- "84_Setpoints_LIT304_Refill_Target_Low"
   TextField "Text field_31" at 1152,339 size 100x22; Text 'RE-FILL'
   IOField "I/O field_44" at 650,299 size 75x22; Authorization "Parameter Change"; FormatPattern 999
      ProcessValue <- "84_Setpoints_LIT304_InitialFill_Target_Low"
   TextField "Text field_32" at 645,272 size 83x22; Text 'Target Low'
   IOField "I/O field_45" at 750,339 size 75x22; Authorization "Parameter Change"; FormatPattern 999
      ProcessValue <- "84_Setpoints_LIT304_Refill_Target"
   TextField "Text field_2" at 100,379 size 220x22; Text 'PIT416 GAS TO DECK PRESS'
   IOField "I/O field_1" at 350,379 size 70x22; FormatPattern 9.9; Unit  Barg
      ProcessValue <- "12_AI_Data_PIT_416_SCALED"
   TextField "Text field_6" at 20,379 size 53x22; Text 'IW810'
   IOField "I/O field_4" at 750,379 size 75x22; Authorization "Parameter Change"; FormatPattern 9.9; Unit  Barg
      ProcessValue <- "84_Setpoints_PIT416_Target"
   TextField "Text field_7" at 100,419 size 220x22; Text 'PIT358 FCW INLET PRESS'
   IOField "I/O field_2" at 350,419 size 70x22; FormatPattern 9.9; Unit  Barg
      ProcessValue <- "12_AI_Data_PIT_358_SCALED"
   IOField "I/O field_3" at 450,419 size 75x22; Authorization "Parameter Change"; FormatPattern 9.9; Unit  Barg
      ProcessValue <- "84_Setpoints_PIT358_InitialFill_LowLow"
   IOField "I/O field_5" at 550,419 size 75x22; Authorization "Parameter Change"; FormatPattern 9.9; Unit  Barg
      ProcessValue <- "84_Setpoints_PIT358_InitialFill_Low"
   IOField "I/O field_6" at 952,419 size 75x22; Authorization "Parameter Change"; FormatPattern 99.9; Unit  Barg
      ProcessValue <- "84_Setpoints_PIT358_InitialFill_High"
   IOField "I/O field_7" at 1052,419 size 75x22; Authorization "Parameter Change"; FormatPattern 99.9; Unit  Barg
      ProcessValue <- "84_Setpoints_PIT358_InitialFill_HighHigh"
   TextField "Text field_8" at 20,419 size 53x22; Text 'IW812'
   TextField "Text field_9" at 1152,419 size 100x22; Text 'INITIAL FILL'
   IOField "I/O field_8" at 450,459 size 75x22; Authorization "Parameter Change"; FormatPattern 9.9; Unit  Barg
      ProcessValue <- "84_Setpoints_PIT358_Refill_LowLow"
   IOField "I/O field_9" at 550,459 size 75x22; Authorization "Parameter Change"; FormatPattern 9.9; Unit  Barg
      ProcessValue <- "84_Setpoints_PIT358_Refill_Low"
   IOField "I/O field_10" at 952,459 size 75x22; Authorization "Parameter Change"; FormatPattern 99.9; Unit  Barg
      ProcessValue <- "84_Setpoints_PIT358_Refill_High"
   IOField "I/O field_11" at 1052,459 size 75x22; Authorization "Parameter Change"; FormatPattern 99.9; Unit  Barg
      ProcessValue <- "84_Setpoints_PIT358_Refill_HighHigh"
   TextField "Text field_10" at 1152,459 size 100x22; Text 'RE-FILL'
   TextField "Text field_3" at 100,499 size 220x22; Text 'PIT353 RECIRC FCW PRESS'
   IOField "I/O field_12" at 350,499 size 70x22; FormatPattern 9.9; Unit  Barg
      ProcessValue <- "12_AI_Data_PIT_353_SCALED"
   IOField "I/O field_13" at 450,499 size 75x22; Authorization "Parameter Change"; FormatPattern 9.9; Unit  Barg
      ProcessValue <- "84_Setpoints_PIT353_InitialFill_LowLow"
   IOField "I/O field_14" at 550,499 size 75x22; Authorization "Parameter Change"; FormatPattern 9.9; Unit  Barg
      ProcessValue <- "84_Setpoints_PIT353_InitialFill_Low"
   IOField "I/O field_15" at 952,499 size 75x22; Authorization "Parameter Change"; FormatPattern 9.9; Unit  Barg
      ProcessValue <- "84_Setpoints_PIT353_InitialFill_High"
   IOField "I/O field_20" at 1052,499 size 75x22; Authorization "Parameter Change"; FormatPattern 9.9; Unit  Barg
      ProcessValue <- "84_Setpoints_PIT353_InitialFill_HighHigh"
   TextField "Text field_4" at 20,499 size 53x22; Text 'IW816'
   TextField "Text field_11" at 1152,499 size 100x22; Text 'INITIAL FILL'
   IOField "I/O field_21" at 450,539 size 75x22; Authorization "Parameter Change"; FormatPattern 9.9; Unit  Barg
      ProcessValue <- "84_Setpoints_PIT353_Refill_LowLow"
   IOField "I/O field_31" at 550,539 size 75x22; Authorization "Parameter Change"; FormatPattern 9.9; Unit  Barg
      ProcessValue <- "84_Setpoints_PIT353_Refill_Low"
   IOField "I/O field_32" at 952,539 size 75x22; Authorization "Parameter Change"; FormatPattern 9.9; Unit  Barg
      ProcessValue <- "84_Setpoints_PIT353_Refill_High"
   IOField "I/O field_33" at 1052,539 size 75x22; Authorization "Parameter Change"; FormatPattern 9.9; Unit  Barg
      ProcessValue <- "84_Setpoints_PIT353_Refill_HighHigh"
   TextField "Text field_12" at 1152,539 size 100x22; Text 'RE-FILL'
   TextField "Text field_5" at 836,272 size 107x22; Text 'Safe Target'
   IOField "I/O field_16" at 854,379 size 75x22; Authorization "Parameter Change"; FormatPattern 9.99; Unit  Barg
      ProcessValue <- "84_Setpoints_PIT416_Target_Safe"
   Group "Group" at 455,41 size 373x50
   Button "HmiScreenItemData_8" at 469,45 size 355x40; TextOn 'Back'; TextOff 'Text'
   TextField "Screen title" at 455,41 size 373x50; Text 'Screen title'

screen "Commissioning Main Page" 1280x800, template "Template"
   on GenerateScreen: "TitleUpdater"()
   Button "HmiScreenItemData_1" at 1,1 size 150x43; TextOn 'Back'; TextOff 'Main Index'
      on Release: ActivateScreen("02 Main Index", 0)
   AlarmView "Alarm view_1" at 0,777 size 1280x23
   Button "HmiScreenItemData_4" at 790,100 size 200x35; TextOn 'Back'; TextOff 'BWT Settings'
   Button "Button_22" at 800,150 size 180x50; TextOff 'Target Setpoints'; Authorization "Commissioning"
      on Press: ActivateScreen("BWT Target Setpoints", 0)
   Button "Button_24" at 800,220 size 180x50; TextOff 'Process Times'; Authorization "Commissioning"
      on Press: ActivateScreen("BWT Process Times", 0)
   Button "HmiScreenItemData_3" at 540,100 size 200x35; TextOn 'Back'; TextOff 'GCU Settings'
   Button "Button_13" at 550,150 size 180x50; TextOff 'Digital Inputs'; Authorization "Commissioning"
      on Click: ActivateScreen("GCU Digital Inputs", 0)
   Button "Button_14" at 550,220 size 180x50; TextOff 'Digital Outputs'; Authorization "Operating Mode"
      on Click: ActivateScreen("GCU Digital Outputs", 0)
   Button "Button_15" at 550,290 size 180x50; TextOff 'Analogue Inputs'; Authorization "Commissioning"
      on Press: ActivateScreen("GCU Analogue Inputs", 0)
   Button "Button_16" at 550,430 size 180x50; TextOff 'Target Setpoints'; Authorization "Commissioning"
      on Press: ActivateScreen("GCU Target Setpoints", 0)
   Button "Button_17" at 550,360 size 180x50; TextOff 'Analogue Outputs'; Authorization "Commissioning"
      on Press: ActivateScreen("GCU Analogue Outputs", 0)
   Button "Button_18" at 550,500 size 180x50; TextOff 'Process Times'; Authorization "Commissioning"
      on Press: ActivateScreen("GCU Process Times", 0)
   Button "HmiScreenItemData_2" at 290,100 size 200x35; TextOn 'Back'; TextOff 'IGG Settings'
   Button "Button_7" at 300,150 size 180x50; TextOff 'Digital Inputs'; Authorization "Commissioning"
      on Click: ActivateScreen("IGG Digital Inputs", 0)
   Button "Button_8" at 300,220 size 180x50; TextOff 'Digital Outputs'; Authorization "Operating Mode"
      on Click: ActivateScreen("IGG Digital Outputs", 0)
   Button "Button_9" at 300,290 size 180x50; TextOff 'Analogue Inputs'; Authorization "Commissioning"
      on Press: ActivateScreen("IGG Analogue Inputs", 0)
   Button "Button_10" at 300,430 size 180x50; TextOff 'Target Setpoints'; Authorization "Commissioning"
      on Press: ActivateScreen("IGG Target Setpoints", 0)
   Button "Button_11" at 300,360 size 180x50; TextOff 'Analogue Outputs'; Authorization "Commissioning"
      on Press: ActivateScreen("IGG Analogue Outputs", 0)
   Button "Button_12" at 300,500 size 180x50; TextOff 'Process Times'; Authorization "Commissioning"
      on Press: ActivateScreen("IGG Process Times", 0)
   Button "HmiScreenItemData_6" at 40,100 size 200x35; TextOn 'Back'; TextOff 'BC Settings'
   Button "Button_1" at 50,150 size 180x50; TextOff 'Digital Inputs'; Authorization "Commissioning"
      on Click: ActivateScreen("BC Digital Inputs", 0)
   Button "Button_2" at 50,220 size 180x50; TextOff 'Digital Outputs'; Authorization "Operating Mode"
      on Click: ActivateScreen("BC Digital Outputs", 0)
   Button "Button_3" at 50,290 size 180x50; TextOff 'Analogue Inputs'; Authorization "Commissioning"
      on Press: ActivateScreen("BC Analogue Inputs", 0)
   Button "Button_5" at 50,430 size 180x50; TextOff 'Target Setpoints'; Authorization "Commissioning"
      on Press: ActivateScreen("BC Target Setpoints", 0)
   Button "Button_4" at 50,360 size 180x50; TextOff 'Analogue Outputs'; Authorization "Commissioning"
      on Press: ActivateScreen("BC Analogue Outputs", 0)
   Button "Button_6" at 50,570 size 180x50; TextOff 'Max Step Times'; Authorization "Commissioning"
      on Press: ActivateScreen("BC Max Step Times", 0)
   Button "HmiScreenItemData_5" at 1040,100 size 200x35; TextOn 'Back'; TextOff 'RIO Racks'
   Button "Button_25" at 1050,150 size 180x32; TextOff 'RIO 1 Digital Inputs'; Authorization "Commissioning"
      on Click: ActivateScreen("RIO 01 Digital Inputs", 0)
   Button "Button_26" at 1050,220 size 180x32; TextOff 'RIO 2 Digital Inputs'; Authorization "Operating Mode"
      on Click: ActivateScreen("RIO 02 Digital Inputs", 0)
   Button "Button_27" at 1050,290 size 180x32; TextOff 'RIO 3 Digital Inputs'; Authorization "Commissioning"
      on Click: ActivateScreen("RIO 03 Digital Inputs", 0)
   Button "Button_28" at 1050,430 size 180x32; TextOff 'RIO 5 Digital Inputs'; Authorization "Commissioning"
      on Click: ActivateScreen("RIO 05 Digital Inputs", 0)
   Button "Button_29" at 1050,360 size 180x32; TextOff 'RIO 4 Digital Inputs'; Authorization "Commissioning"
      on Click: ActivateScreen("RIO 04 Digital Inputs", 0)
   Button "Button_30" at 1050,500 size 180x32; TextOff 'RIO 6 Digital Inputs'; Authorization "Commissioning"
      on Click: ActivateScreen("RIO 06 Digital Inputs", 0)
   Button "Button_31" at 1050,570 size 180x32; TextOff 'RIO 7 Digital Inputs'; Authorization "Commissioning"
      on Click: ActivateScreen("RIO 07 Digital Inputs", 0)